REGION Network 5: Compare
         L     7;
   COMP: NOP   0;
         T     #Loop2;
         L     B[AR1, P#1.0];
         L     B[AR2, P#1.0];
         <I;
         JC    RESE;
         >I;
         JC    SET;
         +AR1  P#1.0;
         +AR2  P#1.0;
         L     #Loop2;
         LOOP  COMP;
   RESE: NOP   0;
         R     #"#COMP_DATETIME";
         JU    END;
   SET:  NOP   0;
         S     #"#COMP_DATETIME";
         JU    END;
END_REGION

REGION Network 6: Error
         JU    ERR;
   ERR:  NOP   0;
         CLR;
         SAVE;
END_REGION

REGION Network 7: End
         JU    END;
   END:  NOP   0;
         L     #SaveSTW;
         T     STW;
         BE;
END_REGION
END_FUNCTION

FUNCTION "#DATA_INPUT_FILTER_EAN13" : Void   // FC306, SCL
TITLE = Data input filter EAN13
{ S7_Optimized_Access := 'FALSE' }
AUTHOR : QLR
FAMILY : dnomaiD
VERSION : 9.0
BEGIN
   #OK := FALSE;
   FOR #"Counter" := #ArrayIni TO #ArrayEnd DO //#Data #OK
       IF (#Data[#"Counter"]>=#Chr_0 AND #Data[#"Counter"]<=#Chr_9) OR #Data[#"Counter"]=#Chr_Space OR #Data[#"Counter"]=#Chr_Null  THEN
           #OK := TRUE;
       ELSE
           #OK := FALSE;
           EXIT;
       END_IF;
   END_FOR;
END_FUNCTION

FUNCTION "#DATA_INPUT_FILTER_HMI_EAN13" : Void   // FC307, SCL
TITLE = Data input filter HMI EAN13
{ S7_Optimized_Access := 'FALSE' }
AUTHOR : QLR
FAMILY : dnomaiD
VERSION : 9.0
BEGIN

   "#DATA_INPUT_FILTER_EAN13"(OK=>#OK, Data:=#Data);

   #ChrSpaceCounter := #ArrayIni;
   FOR #"Counter" := #ArrayIni TO #ArrayEnd DO //Chr Space Counter
       IF (#Data[#"Counter"] = #Chr_Space OR #Data[#"Counter"]=#Chr_Null) AND #OK THEN
           #ChrSpaceCounter := 1 + #ChrSpaceCounter;
       END_IF;
   END_FOR;
   #ChrShift := #ChrSpaceCounter;
   FOR #"Counter" := #ArrayIni TO #ArrayEnd DO //Chr Shift 
       IF (#ChrShift<=#ArrayEnd) AND #OK THEN
           IF #Data[#ChrShift] = #Chr_Null THEN
               #Data[#ChrShift] := #Data[#"Counter"];
               #Data[#"Counter"] := #Chr_Space;
           END_IF;
           #ChrShift := 1 + #ChrShift;
       ELSE
           #"Counter" := #ArrayEnd;
           EXIT;
       END_IF;
   END_FOR;
   FOR #"Counter" := #ArrayIni TO #ArrayEnd DO //Replace Chr_0
       IF (#Data[#"Counter"] = #Chr_Space OR #Data[#"Counter"] = #Chr_Null) AND #OK THEN
           #Data[#"Counter"] := #Chr_0;
       END_IF;
   END_FOR;
END_FUNCTION

ORGANIZATION_BLOCK "Main"   // OB1, LAD, ProgramCycle
TITLE = "Main Program Sweep (Cycle)"
{ S7_Optimized_Access := 'FALSE' }
AUTHOR : QLR
FAMILY : dnomaiD
VERSION : 9.0
BEGIN

REGION Network 1: Data Global
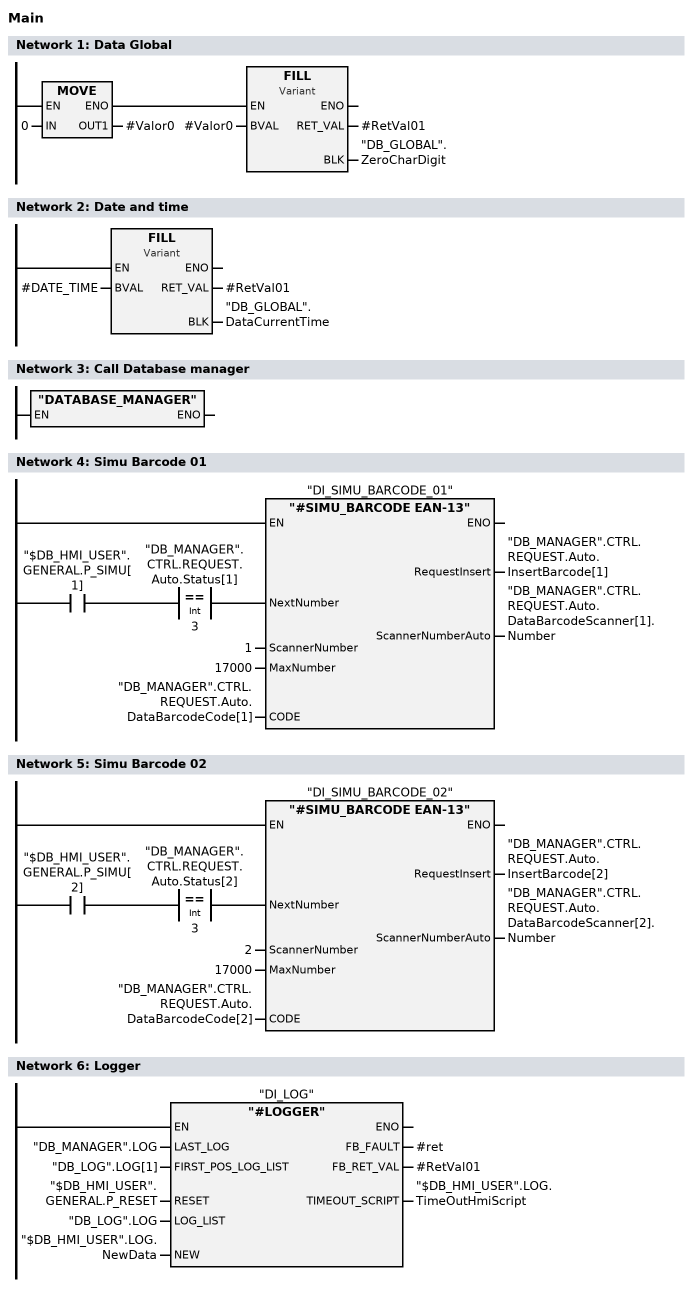
   // ENO of a box is taken as its EN; it also drops when the box reports an error
   #Valor0 := 0;
   #RetVal01 := FILL(BVAL := #Valor0, BLK => "DB_GLOBAL".ZeroCharDigit);
END_REGION

REGION Network 2: Date and time
   #RetVal01 := FILL(BVAL := #DATE_TIME, BLK => "DB_GLOBAL".DataCurrentTime);
END_REGION

REGION Network 3: Call Database manager
   RUNG wire#powerrail
      "DATABASE_MANAGER"()
   END_RUNG
   // the same network as SCL:
   "DATABASE_MANAGER"();
END_REGION

REGION Network 4: Simu Barcode 01
   RUNG wire#powerrail
      "DI_SIMU_BARCODE_01"(NextNumber := wire#w1, ScannerNumber := 1, MaxNumber := 17000, CODE := "DB_MANAGER".CTRL.REQUEST.Auto.DataBarcodeCode[1], RequestInsert => "DB_MANAGER".CTRL.REQUEST.Auto.InsertBarcode[1], ScannerNumberAuto => "DB_MANAGER".CTRL.REQUEST.Auto.DataBarcodeScanner[1].Number)
   END_RUNG
   RUNG wire#powerrail
      Contact( "$DB_HMI_USER".GENERAL.P_SIMU[1] )
      { S7_Templates := "SrcType := Int" } EQ_Contact(in1 := "DB_MANAGER".CTRL.REQUEST.Auto.Status[1], in2 := 3)
   END_RUNG wire#w1
   // the same network as SCL:
   "DI_SIMU_BARCODE_01"(NextNumber := "$DB_HMI_USER".GENERAL.P_SIMU[1] AND ("DB_MANAGER".CTRL.REQUEST.Auto.Status[1] = 3),   // "#SIMU_BARCODE EAN-13"
                        ScannerNumber := 1,
                        MaxNumber := 17000,
                        CODE := "DB_MANAGER".CTRL.REQUEST.Auto.DataBarcodeCode[1],
                        RequestInsert => "DB_MANAGER".CTRL.REQUEST.Auto.InsertBarcode[1],
                        ScannerNumberAuto => "DB_MANAGER".CTRL.REQUEST.Auto.DataBarcodeScanner[1].Number);
END_REGION

REGION Network 5: Simu Barcode 02
   RUNG wire#powerrail
      "DI_SIMU_BARCODE_02"(NextNumber := wire#w1, ScannerNumber := 2, MaxNumber := 17000, CODE := "DB_MANAGER".CTRL.REQUEST.Auto.DataBarcodeCode[2], RequestInsert => "DB_MANAGER".CTRL.REQUEST.Auto.InsertBarcode[2], ScannerNumberAuto => "DB_MANAGER".CTRL.REQUEST.Auto.DataBarcodeScanner[2].Number)
   END_RUNG
   RUNG wire#powerrail
      Contact( "$DB_HMI_USER".GENERAL.P_SIMU[2] )
      { S7_Templates := "SrcType := Int" } EQ_Contact(in1 := "DB_MANAGER".CTRL.REQUEST.Auto.Status[2], in2 := 3)
   END_RUNG wire#w1
   // the same network as SCL:
   "DI_SIMU_BARCODE_02"(NextNumber := "$DB_HMI_USER".GENERAL.P_SIMU[2] AND ("DB_MANAGER".CTRL.REQUEST.Auto.Status[2] = 3),   // "#SIMU_BARCODE EAN-13"
                        ScannerNumber := 2,
                        MaxNumber := 17000,
                        CODE := "DB_MANAGER".CTRL.REQUEST.Auto.DataBarcodeCode[2],
                        RequestInsert => "DB_MANAGER".CTRL.REQUEST.Auto.InsertBarcode[2],
                        ScannerNumberAuto => "DB_MANAGER".CTRL.REQUEST.Auto.DataBarcodeScanner[2].Number);
END_REGION

REGION Network 6: Logger
   RUNG wire#powerrail
      "DI_LOG"(LAST_LOG := "DB_MANAGER".LOG, FIRST_POS_LOG_LIST := "DB_LOG".LOG[1], RESET := "$DB_HMI_USER".GENERAL.P_RESET, LOG_LIST := "DB_LOG".LOG, NEW := "$DB_HMI_USER".LOG.NewData, FB_FAULT => #ret, FB_RET_VAL => #RetVal01, TIMEOUT_SCRIPT => "$DB_HMI_USER".LOG.TimeOutHmiScript)
   END_RUNG
   // the same network as SCL:
   "DI_LOG"(LAST_LOG := "DB_MANAGER".LOG,   // "#LOGGER"
            FIRST_POS_LOG_LIST := "DB_LOG".LOG[1],
            RESET := "$DB_HMI_USER".GENERAL.P_RESET,
            LOG_LIST := "DB_LOG".LOG,
            NEW := "$DB_HMI_USER".LOG.NewData,
            FB_FAULT => #ret,
            FB_RET_VAL => #RetVal01,
            TIMEOUT_SCRIPT => "$DB_HMI_USER".LOG.TimeOutHmiScript);
END_REGION

REGION Network 7: End
END_REGION
END_ORGANIZATION_BLOCK

(* ===== HMI "HMI_RT_1" =====
connection "HMI_Conexión_1": ETHERNET, S7_1500_OMS

HMI tags "Tabla de variables estándar"
   "Test" : Bool, internal
   "AlwaysTRUE" : Bool = PLC "AlwaysTRUE", 1 s
   "AlwaysFALSE" : Bool = PLC "AlwaysFALSE", 1 s
   "Error" : WString[10], internal

HMI tags "USER"
   "$DB_HMI_USER_DATA_MANAGEMENT_BBDD_Delete_BarcodeDig_Digit" : Array [0..12] of Char, 1 s
   "$DB_HMI_USER_DATA_MANAGEMENT_BBDD_Delete_Request" : Bool, 1 s
   "$DB_HMI_USER_DATA_MANAGEMENT_BBDD_Insert_BarcodeData_Code_Digit" : Array [0..12] of Char, 1 s
   "$DB_HMI_USER_DATA_MANAGEMENT_BBDD_Insert_Request" : Bool, 1 s
   "$DB_HMI_USER_DATA_MANAGEMENT_BBDD_Query_BarcodeDig_Digit" : Array [0..12] of Char, 1 s
   "$DB_HMI_USER_DATA_MANAGEMENT_BBDD_Query_Request" : Bool, 1 s
   "$DB_HMI_USER_DATA_MANAGEMENT_P_AUTO_EMPTY" : Bool, 1 s
   "$DB_HMI_USER_GENERAL_P_RESET" : Bool, 1 s
   "$DB_HMI_USER_GENERAL_P_RESET_INSERT_DATA" : Bool, 1 s
   "$DB_HMI_USER_GENERAL_P_SIMU{1}" : Bool, 1 s
   "$DB_HMI_USER_GENERAL_P_SIMU{2}" : Bool, 1 s
   "$DB_HMI_USER_LOG_TimeOutHmiScript" : Bool, 1 s

HMI tags "MANAGER"
   "DB_MANAGER_CTRL_REQUEST_Auto_DataBarcodeCode{1}_Digit" : Array [0..12] of Char, 1 s
   "DB_MANAGER_CTRL_REQUEST_Auto_DataBarcodeCode{2}_Digit" : Array [0..12] of Char, 1 s
   "DB_MANAGER_CTRL_REQUEST_Auto_Status{1}" : Int, 100 ms
   "DB_MANAGER_CTRL_REQUEST_Auto_Status{2}" : Int, 100 ms
   "DB_MANAGER_DATA_REQUEST_Insert_BarcodeData_Code_Digit" : Array [0..12] of Char, 1 s
   "DB_MANAGER_DATA_RESPONSE_InsertData_BarcodeData_Code_Digit" : Array [0..12] of Char, 1 s
   "DB_MANAGER_DATA_STATUS_DataError" : Bool, 1 s
   "DB_MANAGER_DATA_STATUS_Fb_Fault" : Bool, 1 s
   "DB_MANAGER_DATA_STATUS_Mem_Full_nDB{1}" : Bool, 2 s
   "DB_MANAGER_DATA_STATUS_Mem_Full_nDB{2}" : Bool, 2 s
   "DB_MANAGER_DATA_STATUS_Mem_Full_nDB{3}" : Bool, 2 s
   "DB_MANAGER_DATA_STATUS_Mem_Full_nDB{4}" : Bool, 2 s
   "DB_MANAGER_DATA_STATUS_Mem_Full_nDB{5}" : Bool, 2 s
   "DB_MANAGER_DATA_STATUS_Mem_Full_nDB{6}" : Bool, 2 s
   "DB_MANAGER_LIST_DB_QuantityDB" : Int, 1 s
   "DB_MANAGER_LOG_DatabaseTable_BarcodeData_Code_Digit" : Array [0..12] of Char, 100 ms
   "DB_MANAGER_LOG_DatabaseTable_BarcodeData_Scanner_Number" : Int, 100 ms
   "DB_MANAGER_LOG_Request" : Int, 1 s

HMI tags "LOG"
   "Log" : Bool, 100 ms
   "LOG_LOG{1}_DatabaseTable_BarcodeData_Code_Digit" : Array [0..12] of Char, 1 s
   "LOG_LOG{1}_DatabaseTable_BarcodeData_Scanner_Number" : Int, 1 s
   "LOG_LOG{1}_DatabaseTable_DateTime" : Date_And_Time, 1 s
   "LOG_LOG{1}_Request" : Int, 1 s
   "LOG_LOG{10}_DatabaseTable_BarcodeData_Code_Digit" : Array [0..12] of Char, 1 s
   "LOG_LOG{10}_DatabaseTable_BarcodeData_Scanner_Number" : Int, 1 s
   "LOG_LOG{10}_DatabaseTable_DateTime" : Date_And_Time, 1 s
   "LOG_LOG{10}_Request" : Int, 1 s
   "LOG_LOG{2}_DatabaseTable_BarcodeData_Code_Digit" : Array [0..12] of Char, 1 s
   "LOG_LOG{2}_DatabaseTable_BarcodeData_Scanner_Number" : Int, 1 s
   "LOG_LOG{2}_DatabaseTable_DateTime" : Date_And_Time, 1 s
   "LOG_LOG{2}_Request" : Int, 1 s
   "LOG_LOG{3}_DatabaseTable_BarcodeData_Code_Digit" : Array [0..12] of Char, 1 s
   "LOG_LOG{3}_DatabaseTable_BarcodeData_Scanner_Number" : Int, 1 s
   "LOG_LOG{3}_DatabaseTable_DateTime" : Date_And_Time, 1 s
   "LOG_LOG{3}_Request" : Int, 1 s
   "LOG_LOG{4}_DatabaseTable_BarcodeData_Code_Digit" : Array [0..12] of Char, 1 s
   "LOG_LOG{4}_DatabaseTable_BarcodeData_Scanner_Number" : Int, 1 s
   "LOG_LOG{4}_DatabaseTable_DateTime" : Date_And_Time, 1 s
   "LOG_LOG{4}_Request" : Int, 1 s
   "LOG_LOG{5}_DatabaseTable_BarcodeData_Code_Digit" : Array [0..12] of Char, 1 s
   "LOG_LOG{5}_DatabaseTable_BarcodeData_Scanner_Number" : Int, 1 s
   "LOG_LOG{5}_DatabaseTable_DateTime" : Date_And_Time, 1 s
   "LOG_LOG{5}_Request" : Int, 1 s
   "LOG_LOG{6}_DatabaseTable_BarcodeData_Code_Digit" : Array [0..12] of Char, 1 s
   "LOG_LOG{6}_DatabaseTable_BarcodeData_Scanner_Number" : Int, 1 s
   "LOG_LOG{6}_DatabaseTable_DateTime" : Date_And_Time, 1 s
   "LOG_LOG{6}_Request" : Int, 1 s
   "LOG_LOG{7}_DatabaseTable_BarcodeData_Code_Digit" : Array [0..12] of Char, 1 s
   "LOG_LOG{7}_DatabaseTable_BarcodeData_Scanner_Number" : Int, 1 s
   "LOG_LOG{7}_DatabaseTable_DateTime" : Date_And_Time, 1 s
   "LOG_LOG{7}_Request" : Int, 1 s
   "LOG_LOG{8}_DatabaseTable_BarcodeData_Code_Digit" : Array [0..12] of Char, 1 s
   "LOG_LOG{8}_DatabaseTable_BarcodeData_Scanner_Number" : Int, 1 s
   "LOG_LOG{8}_DatabaseTable_DateTime" : Date_And_Time, 1 s
   "LOG_LOG{8}_Request" : Int, 1 s
   "LOG_LOG{9}_DatabaseTable_BarcodeData_Code_Digit" : Array [0..12] of Char, 1 s
   "LOG_LOG{9}_DatabaseTable_BarcodeData_Scanner_Number" : Int, 1 s
   "LOG_LOG{9}_DatabaseTable_DateTime" : Date_And_Time, 1 s
   "LOG_LOG{9}_Request" : Int, 1 s

text list "StatusBBDD": 0 ''; 1 ''

graphic list "StatusBBDD": 0 'BBDD_Ready'; 1 'BBDD_Full'

graphic list "Emptying": 0 'Graphic_5'; 1 'Graphic_4'

SlideinScreen "GraphX_Slidein_Right" 102x768
   Button "Button_1" at 8,26 size 86x80
   Button "Button_2" at 8,146 size 86x80
   Button "Button_3" at 8,266 size 86x80
   Button "Button_4" at 10,656 size 86x80
   Button "Button_5" at 10,526 size 86x80
   Button "Button_6" at 8,386 size 86x80

screen "Logger" 1366x768
   GraphicView "Visor de gráficos_2" at 28,58 size 390x334
   Group "Group" at 29,392 size 368x27
   Group "Group_1" at 29,32 size 271x27
   TextField "Campo de texto_31" at 486,94 size 136x27
   TextField "Campo de texto_32" at 486,139 size 35x27
   TextField "Campo de texto_33" at 487,164 size 41x27
   TextField "Campo de texto_34" at 487,188 size 46x27
   TextField "Campo de texto_35" at 487,212 size 85x27
   TextField "Campo de texto_36" at 521,139 size 95x27
   TextField "Campo de texto_37" at 529,163 size 159x27
   TextField "Campo de texto_38" at 534,187 size 137x27
   TextField "Campo de texto_39" at 574,212 size 142x27
   TextField "Campo de texto_40" at 487,115 size 137x27
   ScreenModuleView "Log[]_1" at 28,429 size 880x32
   ScreenModuleView "Log[]_2" at 28,461 size 880x32
   ScreenModuleView "Log[]_3" at 28,493 size 880x32
   ScreenModuleView "Log[]_4" at 28,525 size 880x32
   ScreenModuleView "Log[]_5" at 28,557 size 880x32
   ScreenModuleView "Log[]_6" at 28,589 size 880x32
   ScreenModuleView "Log[]_7" at 28,621 size 880x32
   ScreenModuleView "Log[]_8" at 28,653 size 880x32
   ScreenModuleView "Log[]_9" at 28,685 size 880x32
   ScreenModuleView "Log[]_10" at 28,717 size 880x32
   ScreenModuleView "ResetAlarm_1" at 1107,704 size 241x51
   ScreenModuleView "ResetAlarm_2" at 1107,640 size 249x51
   TextField "Campo de texto_21" at 29,392 size 138x27
   TextField "Campo de texto_22" at 168,392 size 11x27
   TextField "Campo de texto_23" at 178,392 size 18x27
   TextField "Campo de texto_24" at 197,392 size 14x27
   TextField "Campo de texto_25" at 221,392 size 176x27
   TextField "Campo de texto_26" at 29,32 size 138x27
   TextField "Campo de texto_27" at 168,32 size 11x27
   TextField "Campo de texto_28" at 178,32 size 18x27
   TextField "Campo de texto_29" at 197,32 size 14x27
   TextField "Campo de texto_30" at 221,32 size 79x27

screen "Barcode" 1366x768, template "Template_1"
   TextField "Text field_11" at 411,159 size 56x20
   TextField "Text field_10" at 324,159 size 56x20
   TextField "Text field_9" at 236,159 size 56x20
   TextField "Text field_8" at 147,159 size 56x20
   GraphicView "Graphic view_3" at 141,66 size 70x90
   GraphicView "Graphic view_4" at 228,66 size 70x90
   GraphicView "Graphic view_5" at 315,66 size 70x90
   GraphicView "Graphic view_6" at 402,66 size 70x90
   GraphicIOField "Graphic I/O field_2" at 140,66 size 70x90
   GraphicIOField "Graphic I/O field_3" at 228,66 size 70x90
   GraphicIOField "Graphic I/O field_4" at 316,66 size 70x90
   GraphicIOField "Graphic I/O field_5" at 403,66 size 70x90
   TextField "Text field_2" at 152,39 size 48x27
   TextField "Text field_3" at 241,39 size 48x27
   TextField "Text field_4" at 328,39 size 48x27
   TextField "Text field_5" at 414,39 size 48x27
   SymbolicIOField "Symbolic I/O field_2" at 144,155 size 60x32
   SymbolicIOField "Symbolic I/O field_3" at 232,155 size 60x32
   SymbolicIOField "Symbolic I/O field_4" at 320,155 size 60x32
   SymbolicIOField "Symbolic I/O field_5" at 408,155 size 60x32
   Button "Button_2" at 8,8 size 53x51
   IOField "Campo ES_3" at 583,95 size 272x45
   GraphicView "Graphic view_12" at 519,85 size 71x67
   IOField "Campo ES_4" at 860,105 size 136x29
   ScreenModuleView "Barcode_1" at 40,285 size 576x469
   ScreenModuleView "Barcode_2" at 704,285 size 576x469
   ScreenModuleView "ResetAlarm_1" at 531,152 size 241x51
   ScreenModuleView "ResetAlarm_2" at 533,34 size 241x51
   TextField "Text field_7" at 58,160 size 56x20
   GraphicView "Graphic view_2" at 52,67 size 70x90
   GraphicIOField "Graphic I/O field_1" at 51,67 size 70x90
   TextField "Text field_1" at 63,40 size 48x27
   SymbolicIOField "Symbolic I/O field_1" at 56,156 size 60x32

Template "Template_1" 1366x768
   GraphicView "Graphic view_10" at 1073,0 size 292x217
   TextField "Template_Text field_1" at 13,219 size 24x40
   TextField "Template_Text field_2" at 674,219 size 24x40

PopupScreen "Insert" 240x161
   TextField "Text field_1" at 0,0 size 240x33
   IOField "Campo ES_2" at 6,45 size 227x44
   Button "Botón_1" at 137,115 size 96x32
   Button "Botón_2" at 8,115 size 96x32
   Button "Botón_3" at 208,5 size 22x22

PopupScreen "Delete" 240x161
   TextField "Text field_1" at 0,0 size 240x33
   IOField "Campo ES_2" at 6,45 size 227x44
   Button "Botón_1" at 137,115 size 96x32
   Button "Botón_2" at 8,115 size 96x32
   Button "Botón_3" at 208,5 size 22x22

PopupScreen "Query" 240x161
   TextField "Text field_1" at 0,0 size 240x33
   IOField "Campo ES_2" at 6,45 size 227x44
   Button "Botón_1" at 137,115 size 96x32
   Button "Botón_2" at 8,115 size 96x32
   Button "Botón_3" at 208,5 size 22x22

PopupScreen "Log" 240x161
   TextField "Text field_1" at 0,0 size 240x33
   Button "Botón_3" at 208,5 size 22x22
   Button "Button_6" at 132,56 size 86x80
   Button "Button_1" at 24,56 size 86x80

VB script "Logger"
   Dim file_path, file_name, file, fso, fo, newFile, delimiter, nextLine
   
   'Initialization of Tags
   Const MODE=8	'8 = Append
   delimiter=vbTab
   nextLine=vbCrLf
   newFile = False
   Set fso = CreateObject("Scripting.FilesystemObject")
   file_path = FilePath '"C:\dnomaiD\"
   file_name = "dbms.log"
   file = file_path & file_name
   
   'Start
   If Not NewLog Or Not Enable Or Request <> RequestNumber Then	
   	Logger = False
   	Exit Function
   End If
   
   On Error Resume Next
   
   'Create Folder
   If fso.FolderExists(file_path)  Then
             bfde4b54-0db7-4817-8032-87127bf19bb9 "Path Exist"
       Else 
             fso.CreateFolder (file_path) 
             bfde4b54-0db7-4817-8032-87127bf19bb9 "Path Created"          
   End If 
   If Err.Number<> 0 Then
   	bfde4b54-0db7-4817-8032-87127bf19bb9 "Error # " & CStr(Err.Number)& " "& Err.Description
   	Err.Clear
   	Logger = False	
   	Exit Function
   End If
   
   'Create Text File
   If fso.FileExists(file)  Then
             bfde4b54-0db7-4817-8032-87127bf19bb9 "File Exist"
             newFile = False 
       Else 
             fso.CreateTextFile (file) 
             bfde4b54-0db7-4817-8032-87127bf19bb9 "File Created"          
             newFile = True 
   End If 
   If Err.Number<> 0 Then
   	bfde4b54-0db7-4817-8032-87127bf19bb9 "Error # " & CStr(Err.Number)& " "& Err.Description
   	Err.Clear
   	Logger = False	
   	Exit Function
   End If
   
   'Create a file object
   Set fo= fso.OpenTextFile(file,MODE,True)
   
   'Check if any errors happend
   If Err.Number<> 0 Then
   	bfde4b54-0db7-4817-8032-87127bf19bb9 "Error # " & CStr(Err.Number)& " "& Err.Description
   	Err.Clear
   	Logger = False	
   	Exit Function
   End If
   
   'Write Headline if File is new
   If newFile Then
   	fo.WriteLine("Date" & delimiter & delimiter & delimiter & "Code" & delimiter & delimiter & "Scanner" & nextLine)
   End If
   
   'Write data into file
   fo.WriteLine(Now & delimiter & Code & delimiter & Scanner)
   
   'Close the file
   fo.Close
   
   'Release the Object
   Set fo = Nothing
   Set fso = Nothing
   
   'Return
   Logger = False
   bfde4b54-0db7-4817-8032-87127bf19bb9 "Successful!"

VB script "PowerShellOpenLog"
   Dim fso, File_Path
   Set fso = CreateObject("Wscript.Shell")
   File_Path = FilePath 'C:\Users\Public\dnomaiD\
   
   'Start
   If Not Enable Then
   	bfde4b54-0db7-4817-8032-87127bf19bb9 "Disable"	
   	Exit Sub
   End If
   
   On Error Resume Next
   
   fso.Run("powershell.exe -command Get-Content -Path " & File_Path & "dbms.log -wait;start-sleep 10")
   
   If Err.Number<> 0 Then
   	bfde4b54-0db7-4817-8032-87127bf19bb9 "Error # " & CStr(Err.Number)& " "& Err.Description
   	Err.Clear
   	Exit Sub
   End If
   
   'Release the Object
   Set fso = Nothing

VB script "PowerShellBackup"
   Dim fso, File_Path, DaTi
   Set fso = CreateObject("Wscript.Shell")
   File_Path = FilePath 'C:\Users\Public\dnomaiD\
   DaTi = Year(Now) & Month(Now) & Day(Now) & Hour(Now) & Minute(Now) & Second(Now)
   
   'Start
   If Not Enable Then
   	bfde4b54-0db7-4817-8032-87127bf19bb9 "Disable"	
   	Exit Sub
   End If
   
   On Error Resume Next
   
   fso.Run("powershell.exe -command Rename-Item -Path " & File_Path & "dbms.log " & DaTi & "backup.log;start-sleep 1")
   
   If Err.Number<> 0 Then
   	bfde4b54-0db7-4817-8032-87127bf19bb9 "Error # " & CStr(Err.Number)& " "& Err.Description
   	Err.Clear
   	Exit Sub
   End If
   
   'Release the Object
   Set fso = Nothing
*)

(* ===== HMI "HMI_RT_1" =====

ScreenModuleEditorView "ResetAlarm" 640x480
   Button "Button_1" at 10,10 size 96x51
   GraphicView "Graphic view_8" at 115,10 size 49x51
   TextField "Text field_14" at 174,20 size 101x23
*)

(* ===== HMI "HMI_RT_1" =====

text list "Request": 0 ''; 1 ''; 2 ''; 3 ''; 4 ''; 5 ''; 6 ''

ScreenModuleEditorView "Log[]" 836x44
   IOField "Campo ES_1" at 292,8 size 137x32
   IOField "Campo ES_2" at 604,8 size 26x32
   IOField "Campo ES_3" at 8,8 size 180x32
   TextField "Campo de texto_1" at 186,8 size 112x27
   TextField "Campo de texto_2" at 426,8 size 185x27
   SymbolicIOField "Campo ES simbólico_1" at 637,8 size 251x32
*)

(* ===== HMI "HMI_RT_1" =====

text list "StatusInsertData": 0 ''; 1 ''; 3 ''; 5 ''; 6 ''; 99 ''; 4 ''; 2 ''

graphic list "Simu": 0 'SimuIcon01'; 1 'SimuIcon02'

ScreenModuleEditorView "Barcode" 640x480
   GraphicView "Graphic view_1" at 10,10 size 258x469
   Button "Botón_1" at 80,264 size 65x59
   GraphicView "Visor de gráficos_1" at 238,164 size 333x200
   IOField "Campo ES_1" at 266,326 size 272x45
   SymbolicIOField "Campo ES simbólico_1" at 44,435 size 218x32
   Button "Button_4" at 187,386 size 96x51
   GraphicView "Graphic view_11" at 292,386 size 49x51
*)